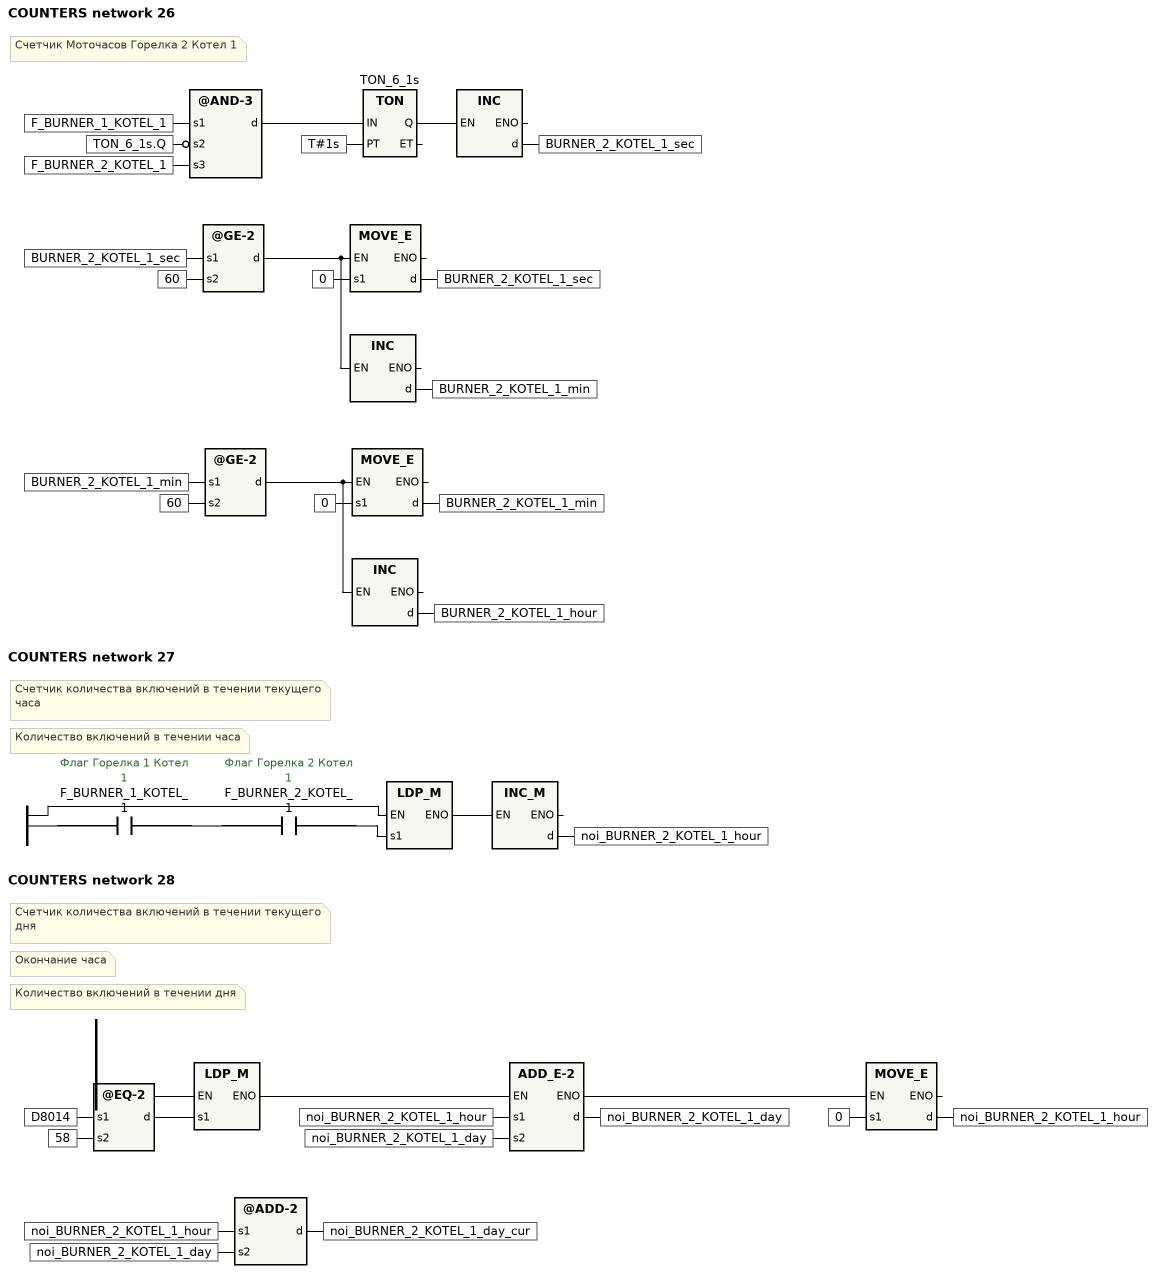
(* [picture p37: structured ladder/FBD of COUNTERS, networks 26 to 28] *)
(* network 26 *)
(* Счетчик Моточасов Горелка 2 Котел 1 *)
TON_6_1s(IN := @AND-3(F_BURNER_1_KOTEL_1, NOT TON_6_1s.Q, F_BURNER_2_KOTEL_1), PT := T#1s);
INC(TON_6_1s.Q, BURNER_2_KOTEL_1_sec);
_p1 := @GE-2(BURNER_2_KOTEL_1_sec, 60);
MOVE_E(_p1, 0, BURNER_2_KOTEL_1_sec);
INC(_p1, BURNER_2_KOTEL_1_min);
_p2 := @GE-2(BURNER_2_KOTEL_1_min, 60);
MOVE_E(_p2, 0, BURNER_2_KOTEL_1_min);
INC(_p2, BURNER_2_KOTEL_1_hour);
(* network 27 *)
(* Счетчик количества включений в течении текущего часа *)
(* Количество включений в течении часа *)
_e1 := LDP_M(TRUE, F_BURNER_1_KOTEL_1 AND F_BURNER_2_KOTEL_1);
INC_M(_e1, noi_BURNER_2_KOTEL_1_hour);
(* network 28 *)
(* Счетчик количества включений в течении текущего дня *)
(* Окончание часа *)
(* Количество включений в течении дня *)
_e1 := LDP_M(TRUE, @EQ-2(D8014, 58));
_e2 := ADD_E(_e1, noi_BURNER_2_KOTEL_1_hour, noi_BURNER_2_KOTEL_1_day, noi_BURNER_2_KOTEL_1_day);
MOVE_E(_e2, 0, noi_BURNER_2_KOTEL_1_hour);
noi_BURNER_2_KOTEL_1_day_cur := @ADD-2(noi_BURNER_2_KOTEL_1_hour, noi_BURNER_2_KOTEL_1_day);
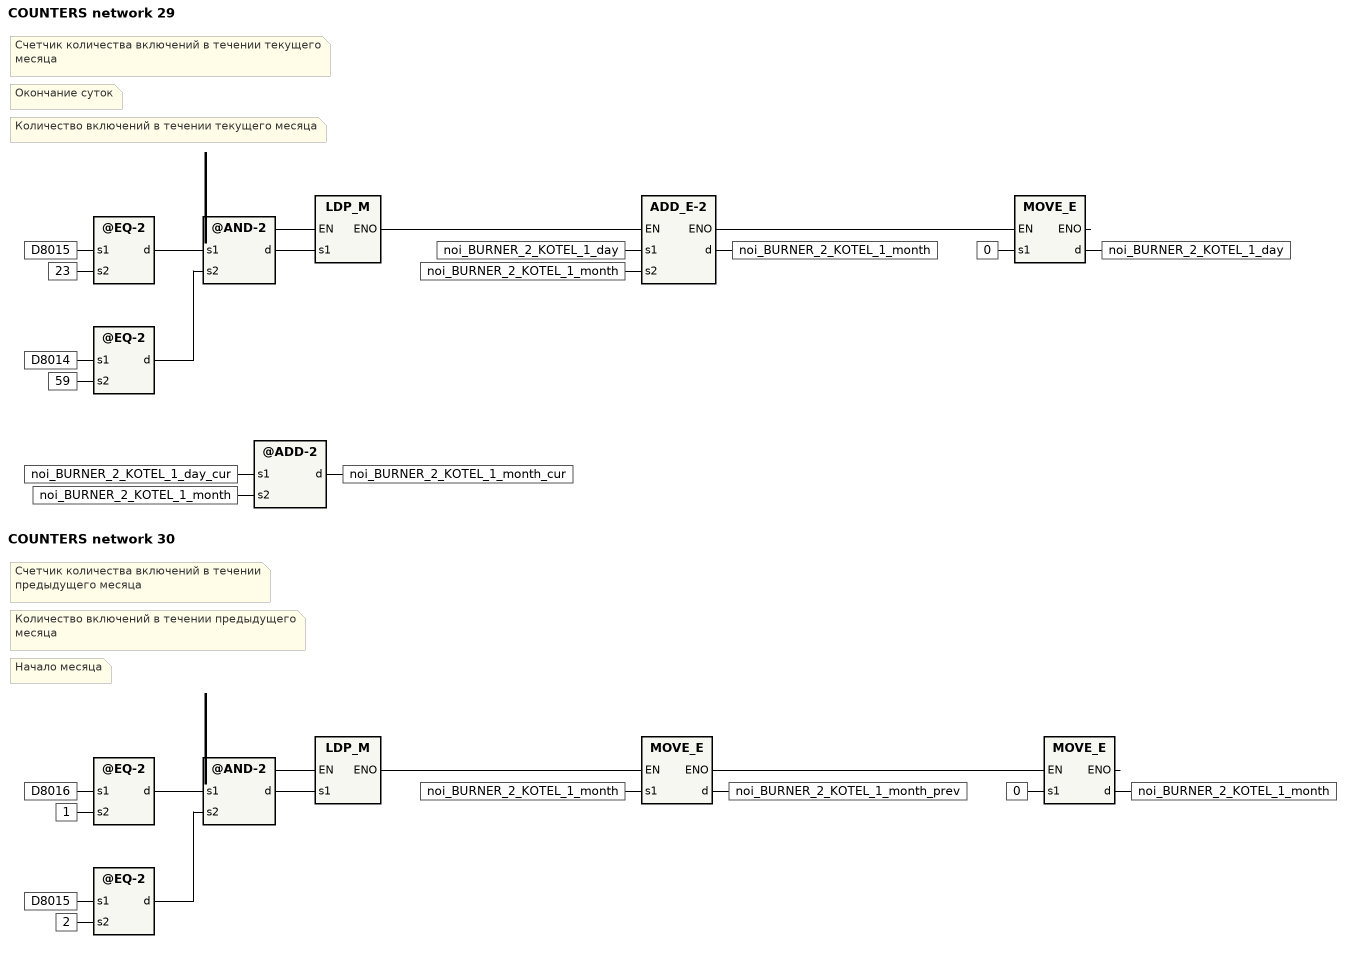
(* network 29 *)
(* Счетчик количества включений в течении текущего месяца *)
(* Окончание суток *)
(* Количество включений в течении текущего месяца *)
_e1 := LDP_M(TRUE, @AND-2(@EQ-2(D8015, 23), @EQ-2(D8014, 59)));
_e2 := ADD_E(_e1, noi_BURNER_2_KOTEL_1_day, noi_BURNER_2_KOTEL_1_month, noi_BURNER_2_KOTEL_1_month);
MOVE_E(_e2, 0, noi_BURNER_2_KOTEL_1_day);
noi_BURNER_2_KOTEL_1_month_cur := @ADD-2(noi_BURNER_2_KOTEL_1_day_cur, noi_BURNER_2_KOTEL_1_month);
(* network 30 *)
(* Счетчик количества включений в течении предыдущего месяца *)
(* Количество включений в течении предыдущего месяца *)
(* Начало месяца *)
_e1 := LDP_M(TRUE, @AND-2(@EQ-2(D8016, 1), @EQ-2(D8015, 2)));
_e2 := MOVE_E(_e1, noi_BURNER_2_KOTEL_1_month, noi_BURNER_2_KOTEL_1_month_prev);
MOVE_E(_e2, 0, noi_BURNER_2_KOTEL_1_month);
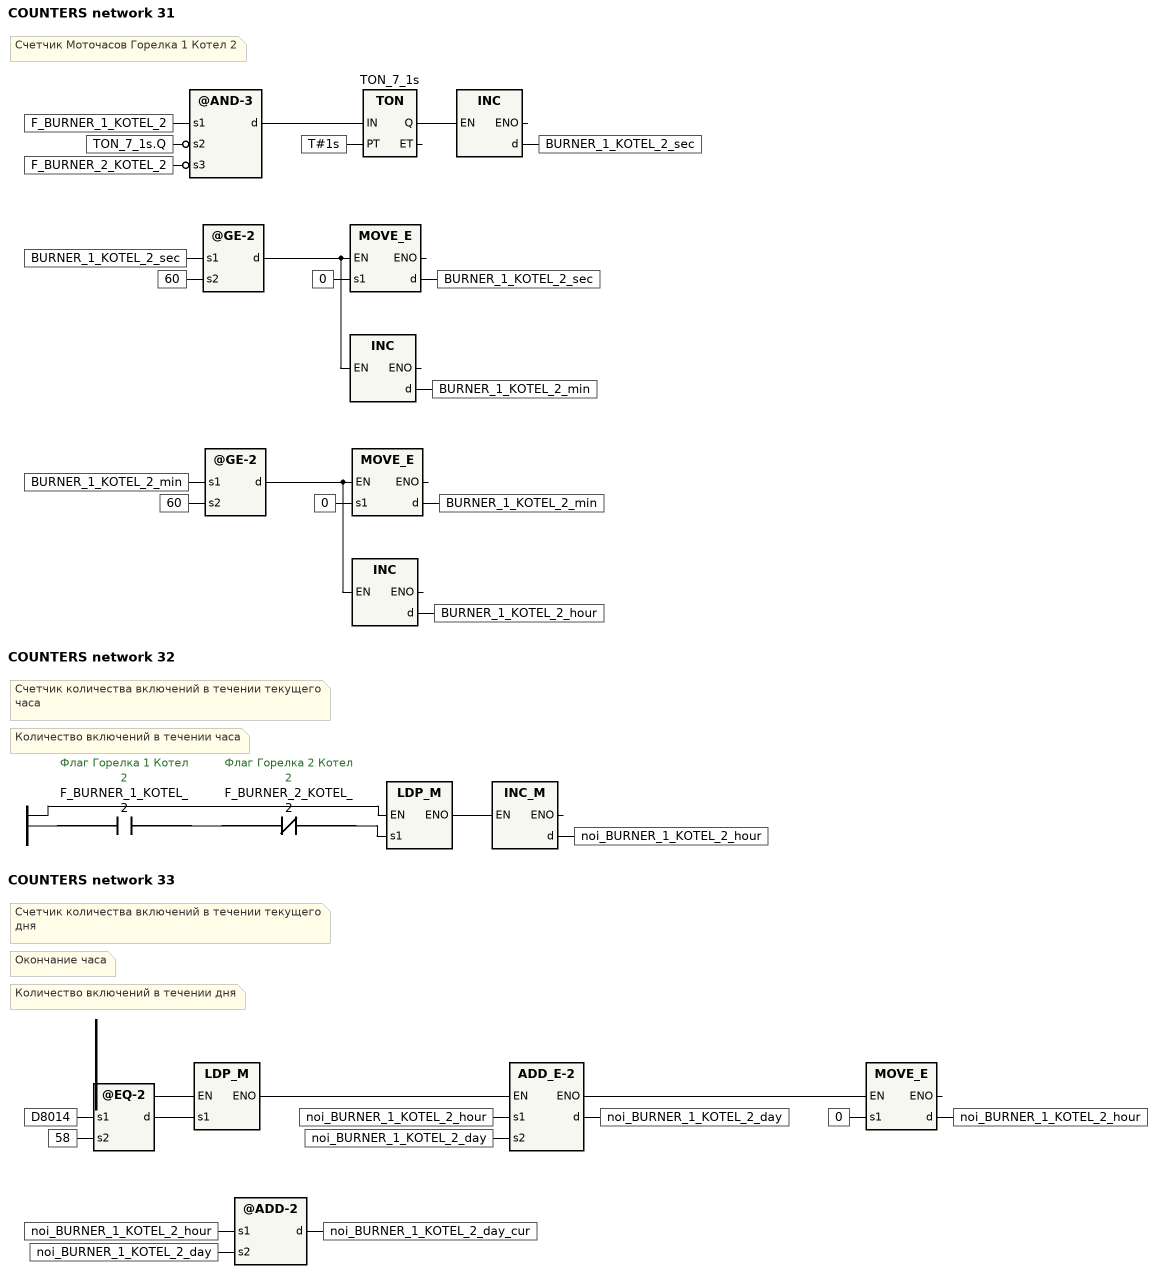
(* network 31 *)
(* Счетчик Моточасов Горелка 1 Котел 2 *)
TON_7_1s(IN := @AND-3(F_BURNER_1_KOTEL_2, NOT TON_7_1s.Q, NOT F_BURNER_2_KOTEL_2), PT := T#1s);
INC(TON_7_1s.Q, BURNER_1_KOTEL_2_sec);
_p1 := @GE-2(BURNER_1_KOTEL_2_sec, 60);
MOVE_E(_p1, 0, BURNER_1_KOTEL_2_sec);
INC(_p1, BURNER_1_KOTEL_2_min);
_p2 := @GE-2(BURNER_1_KOTEL_2_min, 60);
MOVE_E(_p2, 0, BURNER_1_KOTEL_2_min);
INC(_p2, BURNER_1_KOTEL_2_hour);
(* network 32 *)
(* Счетчик количества включений в течении текущего часа *)
(* Количество включений в течении часа *)
_e1 := LDP_M(TRUE, F_BURNER_1_KOTEL_2 AND NOT F_BURNER_2_KOTEL_2);
INC_M(_e1, noi_BURNER_1_KOTEL_2_hour);
(* network 33 *)
(* Счетчик количества включений в течении текущего дня *)
(* Окончание часа *)
(* Количество включений в течении дня *)
_e1 := LDP_M(TRUE, @EQ-2(D8014, 58));
_e2 := ADD_E(_e1, noi_BURNER_1_KOTEL_2_hour, noi_BURNER_1_KOTEL_2_day, noi_BURNER_1_KOTEL_2_day);
MOVE_E(_e2, 0, noi_BURNER_1_KOTEL_2_hour);
noi_BURNER_1_KOTEL_2_day_cur := @ADD-2(noi_BURNER_1_KOTEL_2_hour, noi_BURNER_1_KOTEL_2_day);
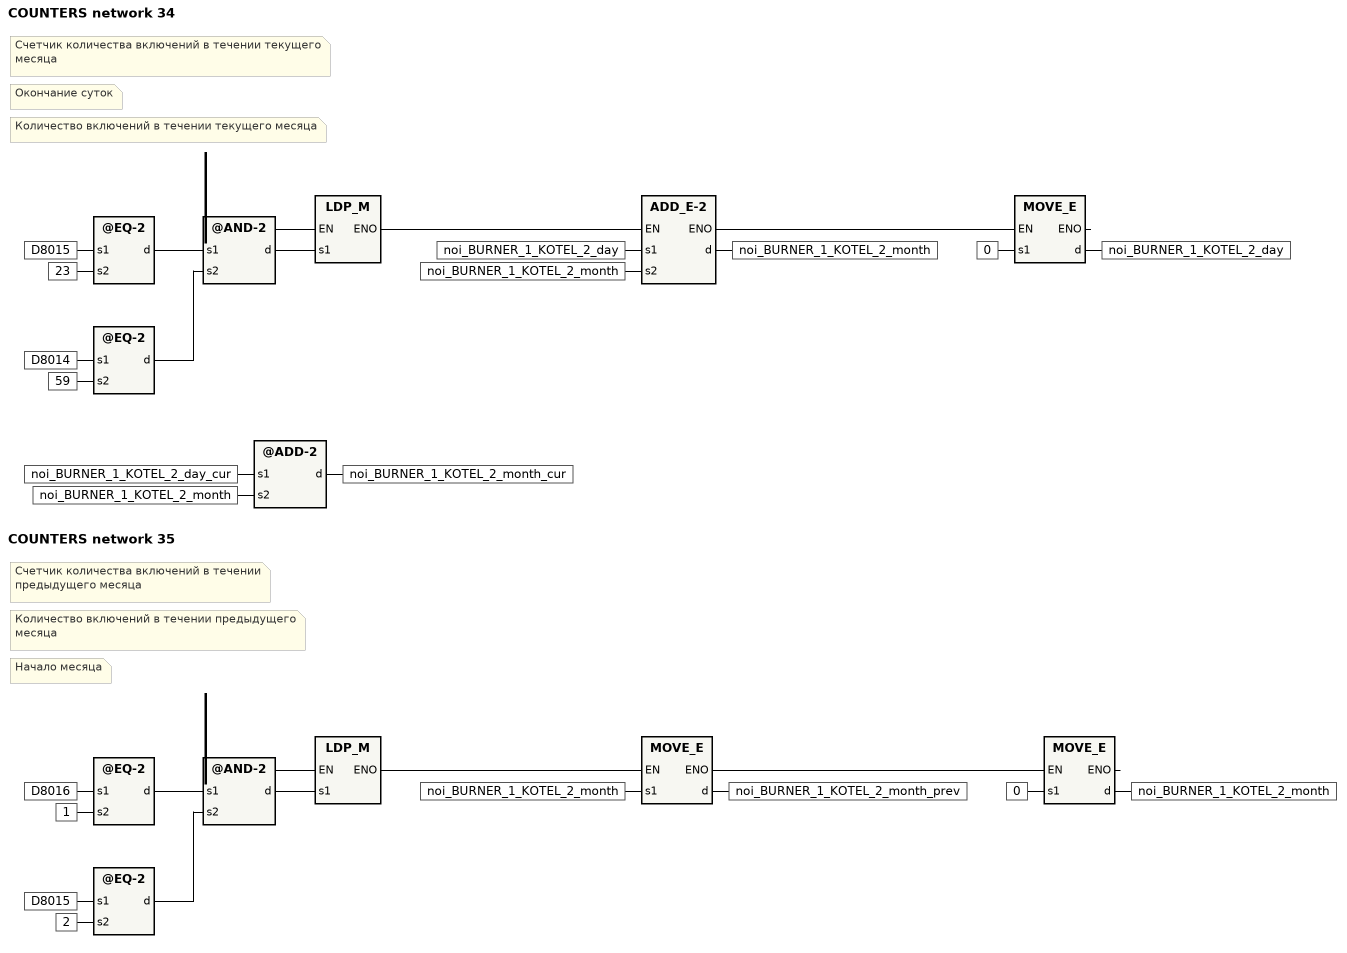
(* network 34 *)
(* Счетчик количества включений в течении текущего месяца *)
(* Окончание суток *)
(* Количество включений в течении текущего месяца *)
_e1 := LDP_M(TRUE, @AND-2(@EQ-2(D8015, 23), @EQ-2(D8014, 59)));
_e2 := ADD_E(_e1, noi_BURNER_1_KOTEL_2_day, noi_BURNER_1_KOTEL_2_month, noi_BURNER_1_KOTEL_2_month);
MOVE_E(_e2, 0, noi_BURNER_1_KOTEL_2_day);
noi_BURNER_1_KOTEL_2_month_cur := @ADD-2(noi_BURNER_1_KOTEL_2_day_cur, noi_BURNER_1_KOTEL_2_month);
(* network 35 *)
(* Счетчик количества включений в течении предыдущего месяца *)
(* Количество включений в течении предыдущего месяца *)
(* Начало месяца *)
_e1 := LDP_M(TRUE, @AND-2(@EQ-2(D8016, 1), @EQ-2(D8015, 2)));
_e2 := MOVE_E(_e1, noi_BURNER_1_KOTEL_2_month, noi_BURNER_1_KOTEL_2_month_prev);
MOVE_E(_e2, 0, noi_BURNER_1_KOTEL_2_month);
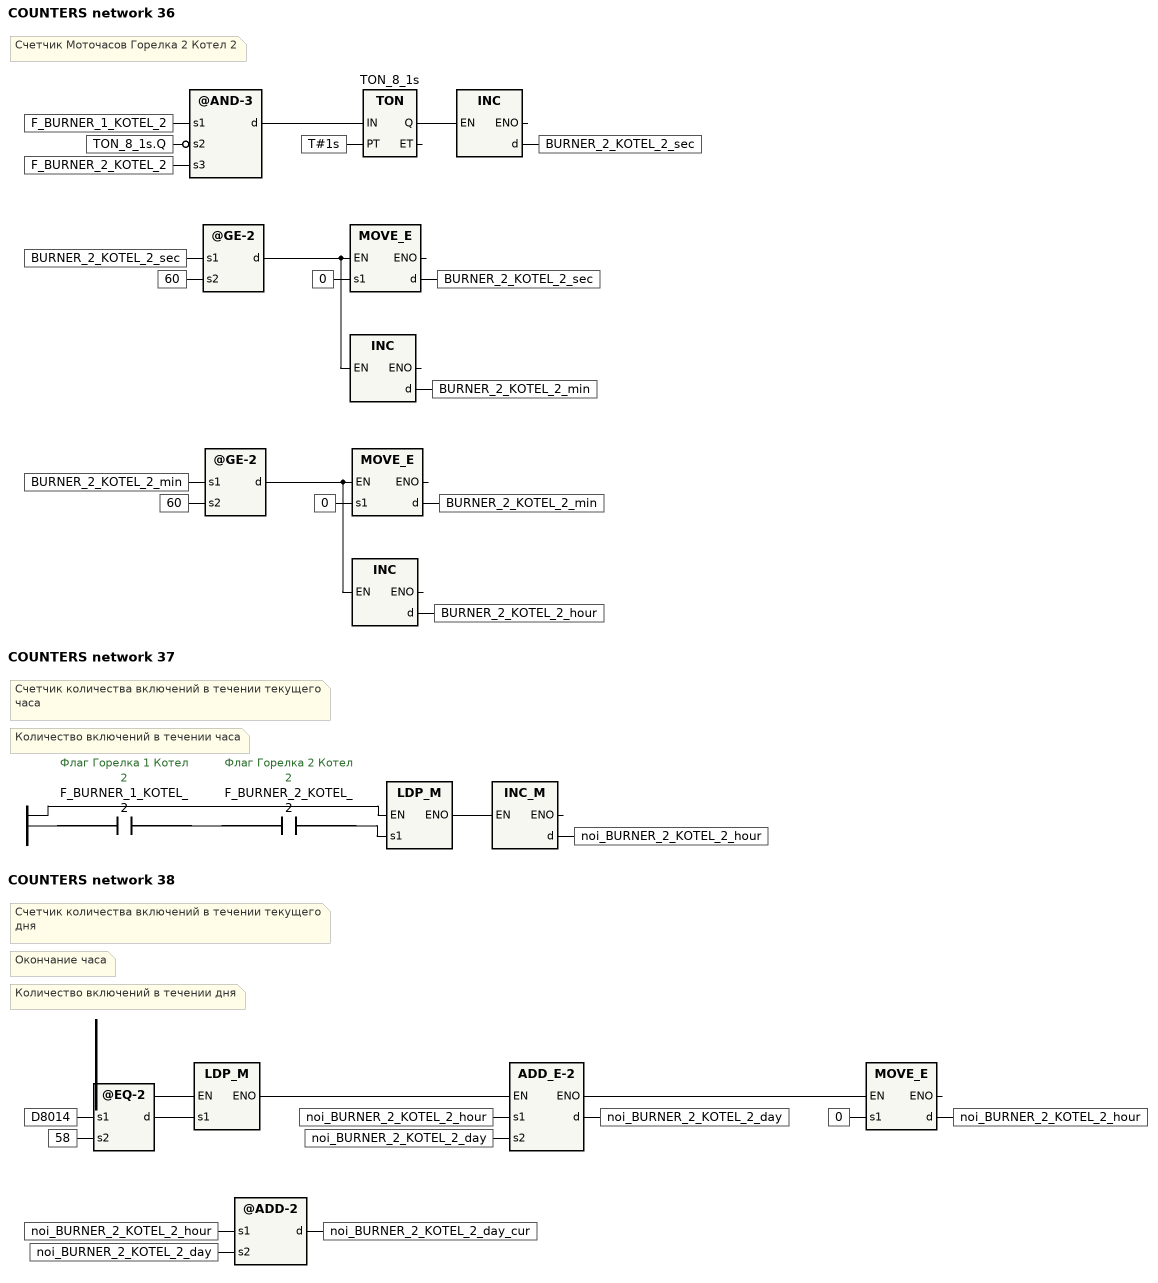
(* network 36 *)
(* Счетчик Моточасов Горелка 2 Котел 2 *)
TON_8_1s(IN := @AND-3(F_BURNER_1_KOTEL_2, NOT TON_8_1s.Q, F_BURNER_2_KOTEL_2), PT := T#1s);
INC(TON_8_1s.Q, BURNER_2_KOTEL_2_sec);
_p1 := @GE-2(BURNER_2_KOTEL_2_sec, 60);
MOVE_E(_p1, 0, BURNER_2_KOTEL_2_sec);
INC(_p1, BURNER_2_KOTEL_2_min);
_p2 := @GE-2(BURNER_2_KOTEL_2_min, 60);
MOVE_E(_p2, 0, BURNER_2_KOTEL_2_min);
INC(_p2, BURNER_2_KOTEL_2_hour);
(* network 37 *)
(* Счетчик количества включений в течении текущего часа *)
(* Количество включений в течении часа *)
_e1 := LDP_M(TRUE, F_BURNER_1_KOTEL_2 AND F_BURNER_2_KOTEL_2);
INC_M(_e1, noi_BURNER_2_KOTEL_2_hour);
(* network 38 *)
(* Счетчик количества включений в течении текущего дня *)
(* Окончание часа *)
(* Количество включений в течении дня *)
_e1 := LDP_M(TRUE, @EQ-2(D8014, 58));
_e2 := ADD_E(_e1, noi_BURNER_2_KOTEL_2_hour, noi_BURNER_2_KOTEL_2_day, noi_BURNER_2_KOTEL_2_day);
MOVE_E(_e2, 0, noi_BURNER_2_KOTEL_2_hour);
noi_BURNER_2_KOTEL_2_day_cur := @ADD-2(noi_BURNER_2_KOTEL_2_hour, noi_BURNER_2_KOTEL_2_day);
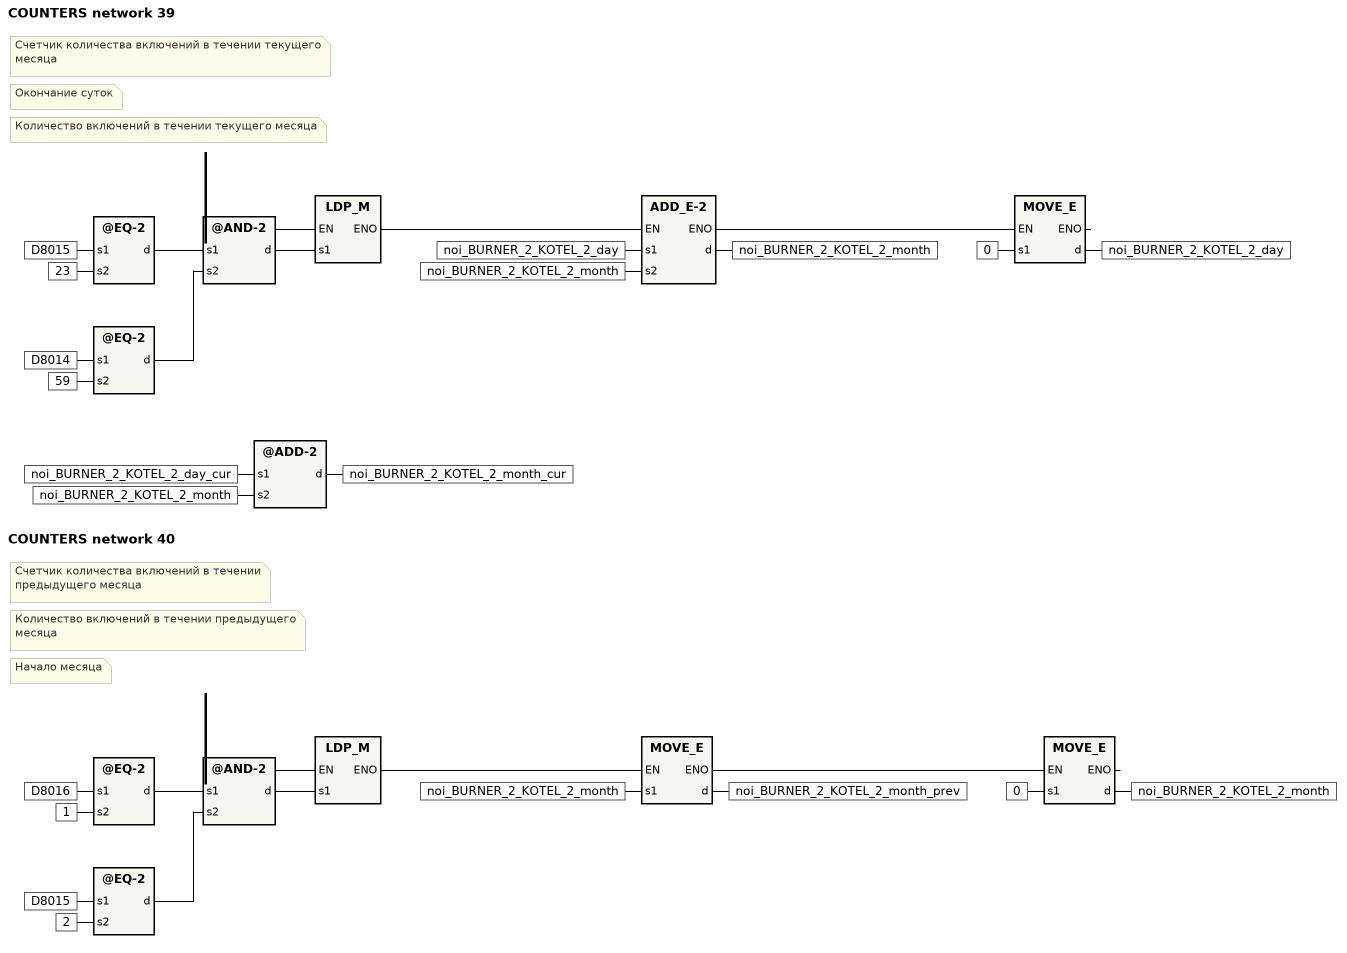
(* network 39 *)
(* Счетчик количества включений в течении текущего месяца *)
(* Окончание суток *)
(* Количество включений в течении текущего месяца *)
_e1 := LDP_M(TRUE, @AND-2(@EQ-2(D8015, 23), @EQ-2(D8014, 59)));
_e2 := ADD_E(_e1, noi_BURNER_2_KOTEL_2_day, noi_BURNER_2_KOTEL_2_month, noi_BURNER_2_KOTEL_2_month);
MOVE_E(_e2, 0, noi_BURNER_2_KOTEL_2_day);
noi_BURNER_2_KOTEL_2_month_cur := @ADD-2(noi_BURNER_2_KOTEL_2_day_cur, noi_BURNER_2_KOTEL_2_month);
(* network 40 *)
(* Счетчик количества включений в течении предыдущего месяца *)
(* Количество включений в течении предыдущего месяца *)
(* Начало месяца *)
_e1 := LDP_M(TRUE, @AND-2(@EQ-2(D8016, 1), @EQ-2(D8015, 2)));
_e2 := MOVE_E(_e1, noi_BURNER_2_KOTEL_2_month, noi_BURNER_2_KOTEL_2_month_prev);
MOVE_E(_e2, 0, noi_BURNER_2_KOTEL_2_month);
END_PROGRAM

PROGRAM EXT_ALARM
(* structured ladder/FBD written out as ST: instructions are called as NAME(EN, inputs, outputs); _pN, _eN, _tN stand for wires *)
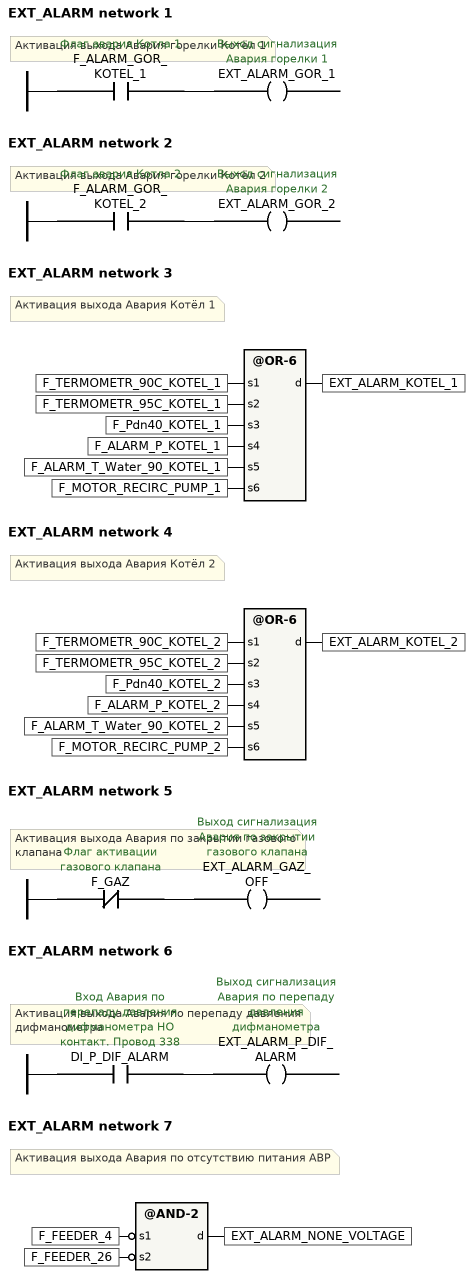
(* network 1 *)
(* Активация выхода Авария горелки Котёл 1 *)
EXT_ALARM_GOR_1 := F_ALARM_GOR_KOTEL_1;
(* network 2 *)
(* Активация выхода Авария горелки Котёл 2 *)
EXT_ALARM_GOR_2 := F_ALARM_GOR_KOTEL_2;
(* network 3 *)
(* Активация выхода Авария Котёл 1 *)
EXT_ALARM_KOTEL_1 := @OR-6(F_TERMOMETR_90C_KOTEL_1, F_TERMOMETR_95C_KOTEL_1, F_Pdn40_KOTEL_1, F_ALARM_P_KOTEL_1, F_ALARM_T_Water_90_KOTEL_1, F_MOTOR_RECIRC_PUMP_1);
(* network 4 *)
(* Активация выхода Авария Котёл 2 *)
EXT_ALARM_KOTEL_2 := @OR-6(F_TERMOMETR_90C_KOTEL_2, F_TERMOMETR_95C_KOTEL_2, F_Pdn40_KOTEL_2, F_ALARM_P_KOTEL_2, F_ALARM_T_Water_90_KOTEL_2, F_MOTOR_RECIRC_PUMP_2);
(* network 5 *)
(* Активация выхода Авария по закрытии газового клапана *)
EXT_ALARM_GAZ_OFF := NOT F_GAZ;
(* network 6 *)
(* Активация выхода Авария по перепаду давления дифманометра *)
EXT_ALARM_P_DIF_ALARM := DI_P_DIF_ALARM;
(* network 7 *)
(* Активация выхода Авария по отсутствию питания АВР *)
EXT_ALARM_NONE_VOLTAGE := @AND-2(NOT F_FEEDER_4, NOT F_FEEDER_26);
END_PROGRAM

PROGRAM FX3UModbusRTUMaster_PRG
VAR
  ModbusComm : FX3UModbusRTUMasterCh2;
  BitOrRegister : BOOL;
  WriteData : ARRAY [0..122] OF WORD;  (* Value of registers to write to slave *)
  CommandCompleted : BOOL;  (* Activates when slave device replies to message *)
  StationNumber : INT;  (* Station no. of slave device *)
  ReadData : ARRAY [0..124] OF WORD;  (* Values read from slave *)
  ReadDataWordCount : INT;
  ReadDataByteCount : INT;
  RegisterStorage : ARRAY [0..124] OF WORD;  (* Values read from slave *)
  BitStorage : ARRAY [0..124] OF WORD;  (* Values read from slave *)
  SequenceCounter : INT;
  Start : BOOL;
  SingleDevices : BOOL;
  ReadOnlyDevices : BOOL;
  StartCommand : BOOL;
  FirstAddress : BOOL;
  ReadOrWrite : BOOL;
  StartAddress : WORD;
  NoOfDevices : INT;
  NoOfReadBits : INT;
  NoOfWriteBits : INT;
  NoOfReadRegisters : INT;
  NoOfWriteRegisters : INT;
  CommandCompletedOk : BOOL;
  CommandCompletedOkCount : INT;
  CommandError : BOOL;  (* Error in communication with slave *)
  CommandErrorCount : INT;
  ResponseTimeoutError : BOOL;
  ResponseTimeoutErrorCount : INT;
  InvalidResponse : BOOL;
  InvalidResponseCount : INT;
  InvalidCommand : BOOL;
  InvalidCommandCount : INT;
  ModbusException : BOOL;
  ModbusExceptionCount : INT;
  ModbusExceptionCode : WORD;
  ModbusExceptionCodeLog : WORD;
  RegisterStorageWater : ARRAY [0..124] OF WORD;  (* Values read from slave *)
END_VAR
(* structured ladder/FBD written out as ST: instructions are called as NAME(EN, inputs, outputs); _pN, _eN, _tN stand for wires *)
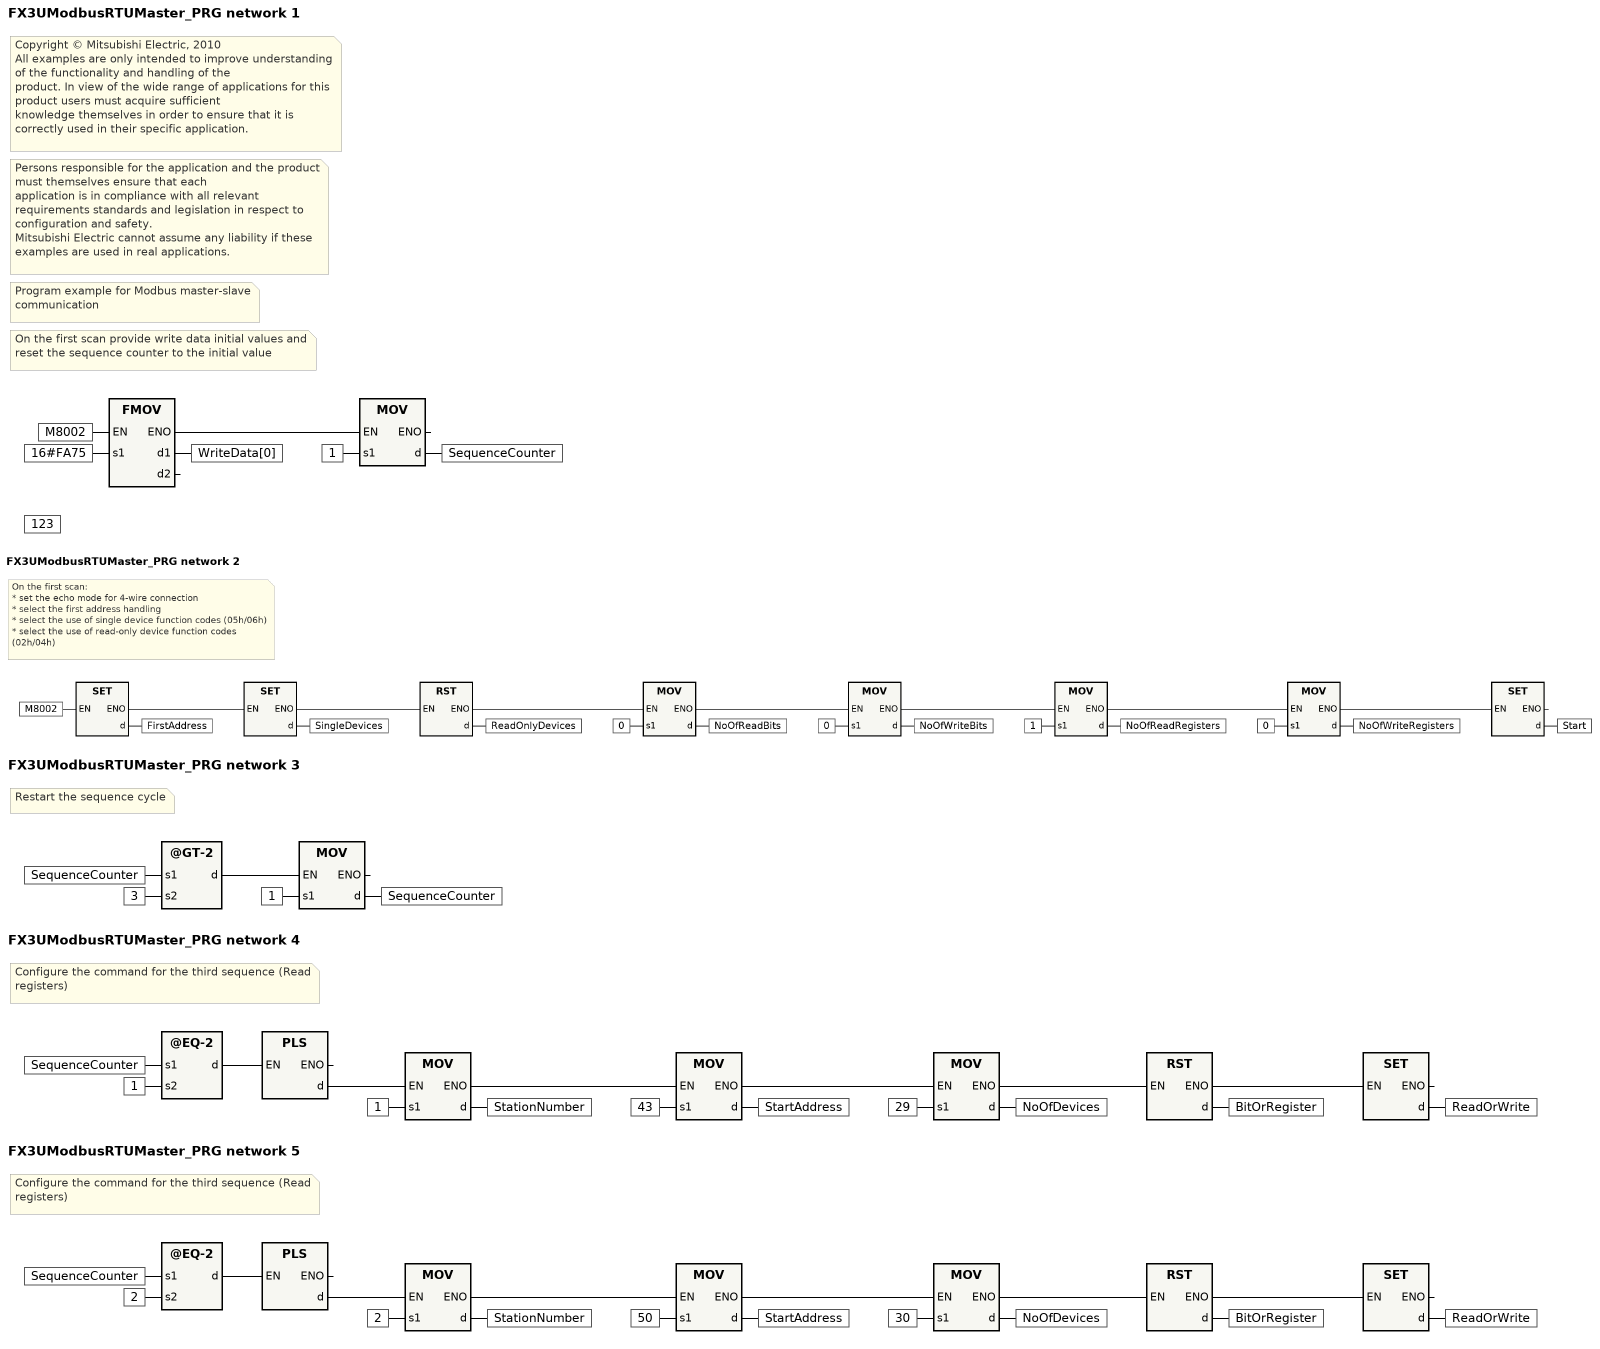
(* network 1 *)
(* Copyright © Mitsubishi Electric, 2010 / All examples are only intended to improve understanding of the functionality and handling of the    / product. In view of the wide range of applications for this product users must acquire sufficient         / knowledge themselves in order to ensure that it is correctly used in their specific application. *)
(* Persons responsible for the application and the product must themselves ensure that each        / application is in compliance with all relevant requirements standards and legislation in respect to    / configuration and safety. /  / Mitsubishi Electric cannot assume any liability if these examples are used in real applications. *)
(* Program example for Modbus master-slave communication *)
(* On the first scan provide write data initial values and reset the sequence counter to the initial value *)
_e1 := FMOV(M8002, 16#FA75, WriteData[0], _open);
MOV(_e1, 1, SequenceCounter);
(* not connected to any output: 123 *)
(* network 2 *)
(* On the first scan:  /  * set the echo mode for 4-wire connection /  * select the first address handling /  * select the use of single device function codes (05h/06h)  /  * select the use of read-only device function codes (02h/04h) *)
_e1 := SET(M8002, FirstAddress);
_e2 := SET(_e1, SingleDevices);
_e3 := RST(_e2, ReadOnlyDevices);
_e4 := MOV(_e3, 0, NoOfReadBits);
_e5 := MOV(_e4, 0, NoOfWriteBits);
_e6 := MOV(_e5, 1, NoOfReadRegisters);
_e7 := MOV(_e6, 0, NoOfWriteRegisters);
SET(_e7, Start);
(* network 3 *)
(* Restart the sequence cycle *)
MOV(@GT-2(SequenceCounter, 3), 1, SequenceCounter);
(* network 4 *)
(* Configure the command for the third sequence (Read registers) *)
PLS(@EQ-2(SequenceCounter, 1), _t1);
_e2 := MOV(_t1, 1, StationNumber);
_e3 := MOV(_e2, 43, StartAddress);
_e4 := MOV(_e3, 29, NoOfDevices);
_e5 := RST(_e4, BitOrRegister);
SET(_e5, ReadOrWrite);
(* network 5 *)
(* Configure the command for the third sequence (Read registers) *)
PLS(@EQ-2(SequenceCounter, 2), _t1);
_e2 := MOV(_t1, 2, StationNumber);
_e3 := MOV(_e2, 50, StartAddress);
_e4 := MOV(_e3, 30, NoOfDevices);
_e5 := RST(_e4, BitOrRegister);
SET(_e5, ReadOrWrite);
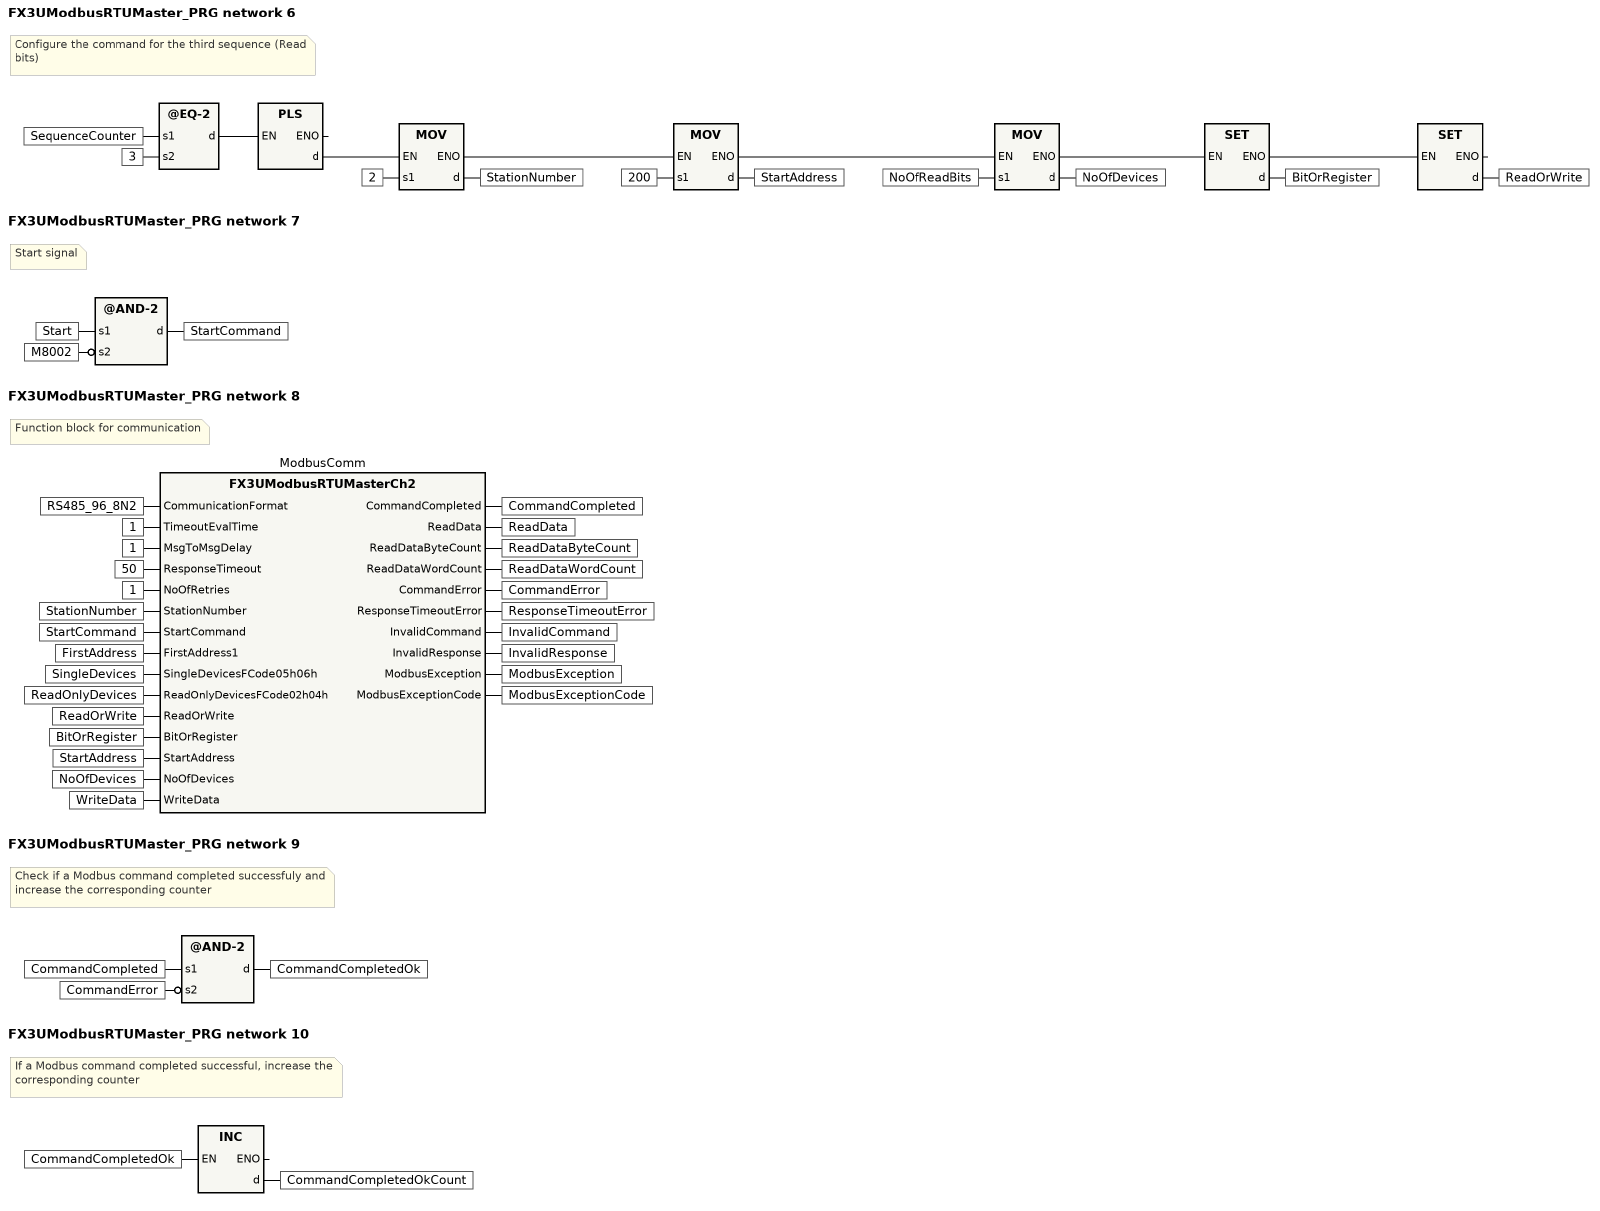
(* network 6 *)
(* Configure the command for the third sequence (Read bits) *)
PLS(@EQ-2(SequenceCounter, 3), _t1);
_e2 := MOV(_t1, 2, StationNumber);
_e3 := MOV(_e2, 200, StartAddress);
_e4 := MOV(_e3, NoOfReadBits, NoOfDevices);
_e5 := SET(_e4, BitOrRegister);
SET(_e5, ReadOrWrite);
(* network 7 *)
(* Start signal *)
StartCommand := @AND-2(Start, NOT M8002);
(* network 8 *)
(* Function block for communication *)
ModbusComm(CommunicationFormat := RS485_96_8N2, TimeoutEvalTime := 1, MsgToMsgDelay := 1, ResponseTimeout := 50, NoOfRetries := 1, StationNumber := StationNumber, StartCommand := StartCommand, FirstAddress1 := FirstAddress, SingleDevicesFCode05h06h := SingleDevices, ReadOnlyDevicesFCode02h04h := ReadOnlyDevices, ReadOrWrite := ReadOrWrite, BitOrRegister := BitOrRegister, StartAddress := StartAddress, NoOfDevices := NoOfDevices, WriteData := WriteData, CommandCompleted => CommandCompleted, ReadData => ReadData, ReadDataByteCount => ReadDataByteCount, ReadDataWordCount => ReadDataWordCount, CommandError => CommandError, ResponseTimeoutError => ResponseTimeoutError, InvalidCommand => InvalidCommand, InvalidResponse => InvalidResponse, ModbusException => ModbusException, ModbusExceptionCode => ModbusExceptionCode);
(* network 9 *)
(* Check if a Modbus command completed successfuly and increase the corresponding counter *)
CommandCompletedOk := @AND-2(CommandCompleted, NOT CommandError);
(* network 10 *)
(* If a Modbus command completed successful, increase the corresponding counter *)
INC(CommandCompletedOk, CommandCompletedOkCount);
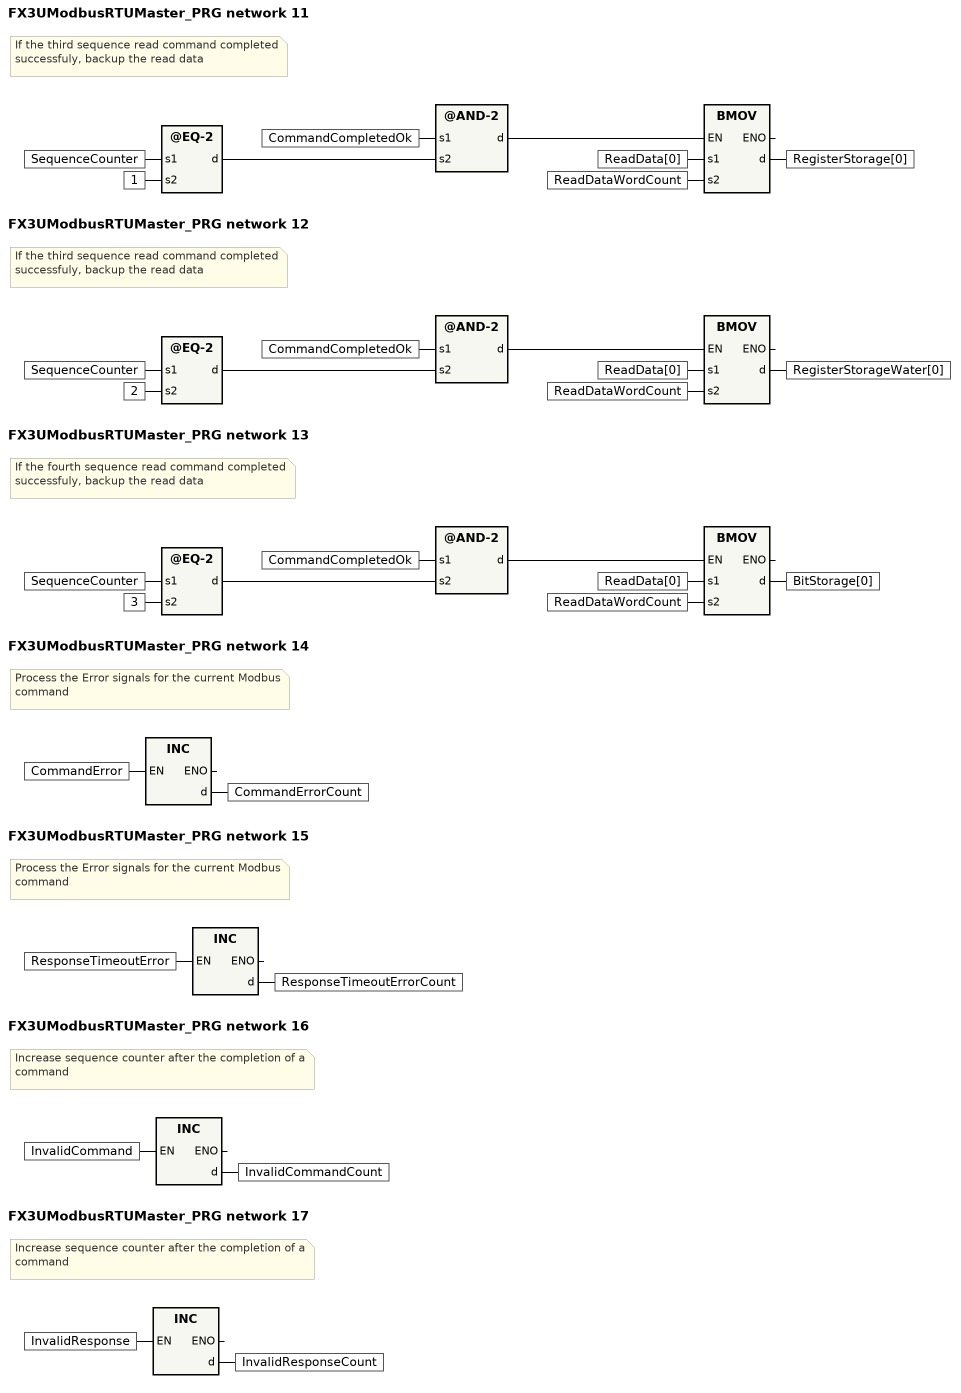
(* network 11 *)
(* If the third sequence read command completed successfuly, backup the read data *)
BMOV(@AND-2(CommandCompletedOk, @EQ-2(SequenceCounter, 1)), ReadData[0], ReadDataWordCount, RegisterStorage[0]);
(* network 12 *)
(* If the third sequence read command completed successfuly, backup the read data *)
BMOV(@AND-2(CommandCompletedOk, @EQ-2(SequenceCounter, 2)), ReadData[0], ReadDataWordCount, RegisterStorageWater[0]);
(* network 13 *)
(* If the fourth sequence read command completed successfuly, backup the read data *)
BMOV(@AND-2(CommandCompletedOk, @EQ-2(SequenceCounter, 3)), ReadData[0], ReadDataWordCount, BitStorage[0]);
(* network 14 *)
(* Process the Error signals for the current Modbus command *)
INC(CommandError, CommandErrorCount);
(* network 15 *)
(* Process the Error signals for the current Modbus command *)
INC(ResponseTimeoutError, ResponseTimeoutErrorCount);
(* network 16 *)
(* Increase sequence counter after the completion of a command *)
INC(InvalidCommand, InvalidCommandCount);
(* network 17 *)
(* Increase sequence counter after the completion of a command *)
INC(InvalidResponse, InvalidResponseCount);
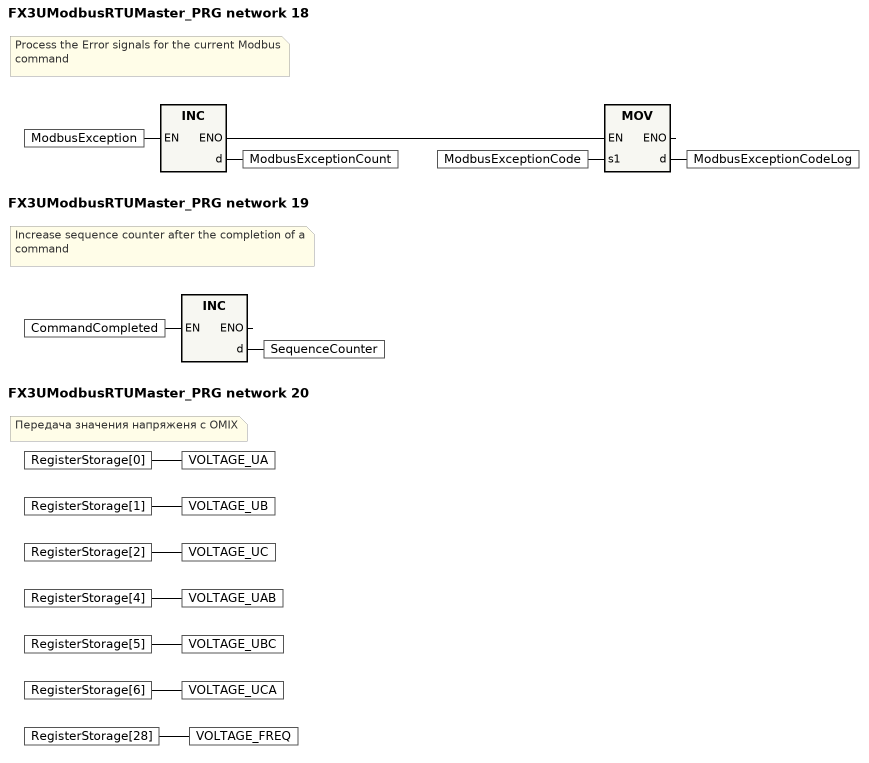
(* network 18 *)
(* Process the Error signals for the current Modbus command *)
_e1 := INC(ModbusException, ModbusExceptionCount);
MOV(_e1, ModbusExceptionCode, ModbusExceptionCodeLog);
(* network 19 *)
(* Increase sequence counter after the completion of a command *)
INC(CommandCompleted, SequenceCounter);
(* network 20 *)
(* Передача значения напряженя с OMIX *)
VOLTAGE_UA := RegisterStorage[0];
VOLTAGE_UB := RegisterStorage[1];
VOLTAGE_UC := RegisterStorage[2];
VOLTAGE_UAB := RegisterStorage[4];
VOLTAGE_UBC := RegisterStorage[5];
VOLTAGE_UCA := RegisterStorage[6];
VOLTAGE_FREQ := RegisterStorage[28];
